// TIA Portal project "EbAndon v4_00_009" (V15) (continued)
DEVICE "ET 200SP station_27"  ET 200SP-Station
   slot 0: "Rack_0"  Rack  6ES5 710-8MAx1
   slot 0: "cv02et200sp"  IM 155-6 PN ST  6ES7 155-6AU01-0BN0  V4.1
   slot 1: "DQ 8x24VDC/0.5A ST_1"  DQ 8x24VDC/0.5A ST  6ES7 132-6BF01-0BA0  V0.0
      slot 1: "DQ 8x24VDC/0.5A ST_1"  DQ 8x24VDC/0.5A ST
   slot 2: "DQ 8x24VDC/0.5A ST_2"  DQ 8x24VDC/0.5A ST  6ES7 132-6BF01-0BA0  V0.0
      slot 1: "DQ 8x24VDC/0.5A ST_2"  DQ 8x24VDC/0.5A ST
   slot 3: "DQ 8x24VDC/0.5A ST_3"  DQ 8x24VDC/0.5A ST  6ES7 132-6BF01-0BA0  V0.0
      slot 1: "DQ 8x24VDC/0.5A ST_3"  DQ 8x24VDC/0.5A ST
   slot 4: "Server module_1"  Server module  6ES7 193-6PA00-0AA0  V1.1
      slot 1: "Server module_1"  Server module
   slot 127: "BA 2xRJ45"  BA 2xRJ45  6ES7 193-6AR00-0AA0  V0.0
      slot 1: "Port_1"  6ES7 193-6AR00-0AA0  V0.0
      slot 2: "Port_2"  6ES7 193-6AR00-0AA0  V0.0
DEVICE "ET 200SP station_28"  ET 200SP-Station
   slot 0: "Rack_0"  Rack  6ES5 710-8MAx1
   slot 0: "cv03et200sp"  IM 155-6 PN ST  6ES7 155-6AU01-0BN0  V4.1
   slot 1: "DQ 8x24VDC/0.5A ST_1"  DQ 8x24VDC/0.5A ST  6ES7 132-6BF01-0BA0  V0.0
      slot 1: "DQ 8x24VDC/0.5A ST_1"  DQ 8x24VDC/0.5A ST
   slot 2: "DQ 8x24VDC/0.5A ST_2"  DQ 8x24VDC/0.5A ST  6ES7 132-6BF01-0BA0  V0.0
      slot 1: "DQ 8x24VDC/0.5A ST_2"  DQ 8x24VDC/0.5A ST
   slot 3: "DQ 8x24VDC/0.5A ST_3"  DQ 8x24VDC/0.5A ST  6ES7 132-6BF01-0BA0  V0.0
      slot 1: "DQ 8x24VDC/0.5A ST_3"  DQ 8x24VDC/0.5A ST
   slot 4: "Server module_1"  Server module  6ES7 193-6PA00-0AA0  V1.1
      slot 1: "Server module_1"  Server module
   slot 127: "BA 2xRJ45"  BA 2xRJ45  6ES7 193-6AR00-0AA0  V0.0
      slot 1: "Port_1"  6ES7 193-6AR00-0AA0  V0.0
      slot 2: "Port_2"  6ES7 193-6AR00-0AA0  V0.0
DEVICE "ET 200SP station_29"  ET 200SP-Station
   slot 0: "Rack_0"  Rack  6ES5 710-8MAx1
   slot 0: "cv04et200sp"  IM 155-6 PN ST  6ES7 155-6AU01-0BN0  V4.1
   slot 1: "DQ 8x24VDC/0.5A ST_1"  DQ 8x24VDC/0.5A ST  6ES7 132-6BF01-0BA0  V0.0
      slot 1: "DQ 8x24VDC/0.5A ST_1"  DQ 8x24VDC/0.5A ST
   slot 2: "DQ 8x24VDC/0.5A ST_2"  DQ 8x24VDC/0.5A ST  6ES7 132-6BF01-0BA0  V0.0
      slot 1: "DQ 8x24VDC/0.5A ST_2"  DQ 8x24VDC/0.5A ST
   slot 3: "DQ 8x24VDC/0.5A ST_3"  DQ 8x24VDC/0.5A ST  6ES7 132-6BF01-0BA0  V0.0
      slot 1: "DQ 8x24VDC/0.5A ST_3"  DQ 8x24VDC/0.5A ST
   slot 4: "Server module_1"  Server module  6ES7 193-6PA00-0AA0  V1.1
      slot 1: "Server module_1"  Server module
   slot 127: "BA 2xRJ45"  BA 2xRJ45  6ES7 193-6AR00-0AA0  V0.0
      slot 1: "Port_1"  6ES7 193-6AR00-0AA0  V0.0
      slot 2: "Port_2"  6ES7 193-6AR00-0AA0  V0.0
DEVICE "ET 200SP station_30"  ET 200SP-Station
   slot 0: "Rack_0"  Rack  6ES5 710-8MAx1
   slot 0: "pc01et200sp"  IM 155-6 PN ST  6ES7 155-6AU01-0BN0  V4.1
   slot 1: "DQ 8x24VDC/0.5A ST_1"  DQ 8x24VDC/0.5A ST  6ES7 132-6BF01-0BA0  V0.0
      slot 1: "DQ 8x24VDC/0.5A ST_1"  DQ 8x24VDC/0.5A ST
   slot 2: "DQ 8x24VDC/0.5A ST_2"  DQ 8x24VDC/0.5A ST  6ES7 132-6BF01-0BA0  V0.0
      slot 1: "DQ 8x24VDC/0.5A ST_2"  DQ 8x24VDC/0.5A ST
   slot 3: "DQ 8x24VDC/0.5A ST_3"  DQ 8x24VDC/0.5A ST  6ES7 132-6BF01-0BA0  V0.0
      slot 1: "DQ 8x24VDC/0.5A ST_3"  DQ 8x24VDC/0.5A ST
   slot 4: "Server module_1"  Server module  6ES7 193-6PA00-0AA0  V1.1
      slot 1: "Server module_1"  Server module
   slot 127: "BA 2xRJ45"  BA 2xRJ45  6ES7 193-6AR00-0AA0  V0.0
      slot 1: "Port_1"  6ES7 193-6AR00-0AA0  V0.0
      slot 2: "Port_2"  6ES7 193-6AR00-0AA0  V0.0
DEVICE "ET 200SP station_31"  ET 200SP-Station
   slot 0: "Rack_0"  Rack  6ES5 710-8MAx1
   slot 0: "pc02et200sp"  IM 155-6 PN ST  6ES7 155-6AU01-0BN0  V4.1
   slot 1: "DQ 8x24VDC/0.5A ST_1"  DQ 8x24VDC/0.5A ST  6ES7 132-6BF01-0BA0  V0.0
      slot 1: "DQ 8x24VDC/0.5A ST_1"  DQ 8x24VDC/0.5A ST
   slot 2: "DQ 8x24VDC/0.5A ST_2"  DQ 8x24VDC/0.5A ST  6ES7 132-6BF01-0BA0  V0.0
      slot 1: "DQ 8x24VDC/0.5A ST_2"  DQ 8x24VDC/0.5A ST
   slot 3: "DQ 8x24VDC/0.5A ST_3"  DQ 8x24VDC/0.5A ST  6ES7 132-6BF01-0BA0  V0.0
      slot 1: "DQ 8x24VDC/0.5A ST_3"  DQ 8x24VDC/0.5A ST
   slot 4: "Server module_1"  Server module  6ES7 193-6PA00-0AA0  V1.1
      slot 1: "Server module_1"  Server module
   slot 127: "BA 2xRJ45"  BA 2xRJ45  6ES7 193-6AR00-0AA0  V0.0
      slot 1: "Port_1"  6ES7 193-6AR00-0AA0  V0.0
      slot 2: "Port_2"  6ES7 193-6AR00-0AA0  V0.0
*)

// ===== PLC "PLC_1"  CPU 1517F-3 PN/DP =====

VAR_GLOBAL   // PLC tag table "Default tag table"
   "System_Byte" AT %MB1 : Byte;
   "FirstScan" AT %M1.0 : Bool;
   "DiagStatUpdt" AT %M1.1 : Bool;
   "AlwaysTRUE" AT %M1.2 : Bool;
   "AlwaysFALSE" AT %M1.3 : Bool;
   "Clock_Byte" AT %MB0 : Byte;
   "Clock_10Hz" AT %M0.0 : Bool;
   "Clock_5Hz" AT %M0.1 : Bool;
   "Clock_2.5Hz" AT %M0.2 : Bool;
   "Clock_2Hz" AT %M0.3 : Bool;
   "Clock_1.25Hz" AT %M0.4 : Bool;
   "Clock_1Hz" AT %M0.5 : Bool;
   "Clock_0.625Hz" AT %M0.6 : Bool;
   "Clock_0.5Hz" AT %M0.7 : Bool;
   "Temp Reset" AT %M2.0 : Bool;
   "clearPartData" AT %M100.0 : Bool;
   "setDefaultPresets" AT %M100.1 : Bool;
   "hardInitReq" AT %M100.2 : Bool;
   "dbg" AT %M500.0 : Bool;
   "dbgSetDefTimes" AT %M5000.0 : Bool;
   "Copy PN Codes Into Recipes" AT %M10.0 : Bool;
   "Load Default Recipes Into Stations" AT %M10.1 : Bool;
   "Load Default Wip Data" AT %M10.2 : Bool;
   "dbg_station_index" AT %MW502 : Int;
END_VAR

VAR_GLOBAL CONSTANT   // PLC tag table "Default tag table"
   "ptsPerStn" : Int := 7;
   "slct_stn_btn_count" : Int := 11;
   "null_value" : Int := -1;
   "wip_pop_up_button_count" : Int := 6;   // number of wip select buttons on wip select pop up screen
END_VAR

VAR_GLOBAL   // PLC tag table "VOLVO 16 01"
   "VOLVO 16 01 IO" AT %QD1000 : DWord;
   "VOLVO 16 01 KP8 In" AT %ID0 : DWord;
   "VOLVO 16 01 KP8 Out" AT %QD0 : DWord;
END_VAR

VAR_GLOBAL   // PLC tag table "VOLVO 16 02"
   "VOLVO 16 02 IO" AT %QD1004 : DWord;
   "VOLVO 16 02 KP8 In" AT %ID4 : DWord;
   "VOLVO 16 02 KP8 Out" AT %QD4 : DWord;
END_VAR

VAR_GLOBAL   // PLC tag table "VOLVO 16 03"
   "VOLVO 16 03 IO" AT %QD1008 : DWord;
   "VOLVO 16 03 KP8 In" AT %ID8 : DWord;
   "VOLVO 16 03 KP8 Out" AT %QD8 : DWord;
END_VAR

VAR_GLOBAL   // PLC tag table "VOLVO 16 04"
   "VOLVO 16 04 IO" AT %QD1012 : DWord;
   "VOLVO 16 04 KP8 In" AT %ID12 : DWord;
   "VOLVO 16 04 KP8 Out" AT %QD12 : DWord;
END_VAR

VAR_GLOBAL   // PLC tag table "VOLVO 16 05"
   "VOLVO 16 05 IO" AT %QD1016 : DWord;
   "VOLVO 16 05 KP8 In" AT %ID16 : DWord;
   "VOLVO 16 05 KP8 Out" AT %QD16 : DWord;
END_VAR

VAR_GLOBAL   // PLC tag table "VOLVO 16 06"
   "VOLVO 16 06 IO" AT %QD1020 : DWord;
   "VOLVO 16 06 KP8 In" AT %ID20 : DWord;
   "VOLVO 16 06 KP8 Out" AT %QD20 : DWord;
END_VAR

VAR_GLOBAL   // PLC tag table "VOLVO 16 07"
   "VOLVO 16 07 IO" AT %QD1024 : DWord;
   "VOLVO 16 07 KP8 In" AT %ID24 : DWord;
   "VOLVO 16 07 KP8 Out" AT %QD24 : DWord;
END_VAR

VAR_GLOBAL   // PLC tag table "VOLVO 16 08"
   "VOLVO 16 08 IO" AT %QD1028 : DWord;
   "VOLVO 16 08 KP8 In" AT %ID28 : DWord;
   "VOLVO 16 08 KP8 Out" AT %QD28 : DWord;
END_VAR

VAR_GLOBAL   // PLC tag table "VOLVO 16 09"
   "VOLVO 16 09 IO" AT %QD1032 : DWord;
   "VOLVO 16 09 KP8 In" AT %ID32 : DWord;
   "VOLVO 16 09 KP8 Out" AT %QD32 : DWord;
END_VAR

VAR_GLOBAL   // PLC tag table "VOLVO 16 10"
   "VOLVO 16 10 IO" AT %QD1036 : DWord;
   "VOLVO 16 10 KP8 In" AT %ID36 : DWord;
   "VOLVO 16 10 KP8 Out" AT %QD36 : DWord;
END_VAR

VAR_GLOBAL   // PLC tag table "VOLVO 16 11"
   "VOLVO 16 11 IO" AT %QD1040 : DWord;
   "VOLVO 16 11 KP8 In" AT %ID40 : DWord;
   "VOLVO 16 11 KP8 Out" AT %QD40 : DWord;
END_VAR

VAR_GLOBAL   // PLC tag table "CHM 02"
   "CHM 02 KP8 In" AT %ID44 : DWord;
   "CHM 02 KP8 Out" AT %QD44 : DWord;
   "CHM 02 IO" AT %QD1044 : DWord;
END_VAR

VAR_GLOBAL   // PLC tag table "CHM 03"
   "CHM 03 IO" AT %QD1048 : DWord;
   "CHM 03 KP8 In" AT %ID48 : DWord;
   "CHM 03 KP8 Out" AT %QD48 : DWord;
END_VAR

VAR_GLOBAL   // PLC tag table "CHM 04"
   "CHM 04 IO" AT %QD1052 : DWord;
   "CHM 04 KP8 In" AT %ID52 : DWord;
   "CHM 04 KP8 Out" AT %QD52 : DWord;
END_VAR

VAR_GLOBAL   // PLC tag table "CHM 05"
   "CHM 05 IO" AT %QD1056 : DWord;
   "CHM 05 KP8 In" AT %ID56 : DWord;
   "CHM 05 KP8 Out" AT %QD56 : DWord;
END_VAR

VAR_GLOBAL   // PLC tag table "CDO 01"
   "CDO 01 IO" AT %QD1060 : DWord;
   "CDO 01 KP8 In" AT %ID60 : DWord;
   "CDO 01 KP8 Out" AT %QD60 : DWord;
END_VAR

VAR_GLOBAL   // PLC tag table "CDO 02"
   "CDO 02 IO" AT %QD1064 : DWord;
   "CDO 02 KP8 In" AT %ID64 : DWord;
   "CDO 02 KP8 Out" AT %QD64 : DWord;
END_VAR

VAR_GLOBAL   // PLC tag table "CDO 03"
   "CDO 03 IO" AT %QD1068 : DWord;
   "CDO 03 KP8 In" AT %ID68 : DWord;
   "CDO 03 KP8 Out" AT %QD68 : DWord;
END_VAR

VAR_GLOBAL   // PLC tag table "BFL 01"
   "BFL 01 IO" AT %QD1072 : DWord;
   "BFL 01 KP8 In" AT %ID72 : DWord;
   "BFL 01 KP8 Out" AT %QD72 : DWord;
   "Manual Operations Trigger" AT %M10.3 : Bool;
END_VAR

VAR_GLOBAL   // PLC tag table "BFL 02"
   "BFL 02 IO" AT %QD1076 : DWord;
   "BFL 02 KP8 In" AT %ID76 : DWord;
   "BFL 02 KP8 Out" AT %QD76 : DWord;
END_VAR

VAR_GLOBAL   // PLC tag table "BFL 03"
   "BFL 03 IO" AT %QD1080 : DWord;
   "BFL 03 KP8 In" AT %ID80 : DWord;
   "BFL 03 KP8 Out" AT %QD80 : DWord;
END_VAR

VAR_GLOBAL   // PLC tag table "LGS 01"
   "LGS 01 IO" AT %QD1084 : DWord;
   "LGS 01 KP8 In" AT %ID84 : DWord;
   "LGS 01 KP8 Out" AT %QD84 : DWord;
END_VAR

VAR_GLOBAL   // PLC tag table "LGS 02"
   "LGS 02 IO" AT %QD1088 : DWord;
   "LGS 02 KP8 In" AT %ID88 : DWord;
   "LGS 02 KP8 Out" AT %QD88 : DWord;
END_VAR

VAR_GLOBAL   // PLC tag table "CHM 01"
   "CHM 01 IO" AT %QD1092 : DWord;
   "CHM 01 KP8 In" AT %ID92 : DWord;
   "CHM 01 KP8 Out" AT %QD92 : DWord;
END_VAR

VAR_GLOBAL CONSTANT   // PLC tag table "Comm Diag"
   "pnioDeviceCount" : Int := 48;   // Upper limit of devices per HMI screen
   "USERDIAG_SLOTS_PER_SCREEN_UPPER_LIM" : Int := 31;   // Upper limit of slots per HMI screen
   "USERDIAG_SLOTS_PER_DEVICE_UPPER_LIM" : Int := 31;   // max number of modules per device
   "USERDIAG_DEVICES_PER_IO_SYSTEM_UPPER_LIM" : Int := 128;   // Upper limit of devices/slaves per IO-System/DP-Mastersystem
   "USERDIAG_SLOTS_PER_PLC_UPPER_LIM" : Int := 31;   // max number of local modules
   "USERDIAG_IO_SYSTEMS_UPPER_LIM" : Int := 1;   // Upper limit of IO-Systems/DP-Mastersystems
   "USERDIAG_IOSYSTEM_1" : Int := 1;   // Index for first IO-System/DP-Mastersystem
END_VAR

VAR_GLOBAL CONSTANT   // PLC tag table "Color Library"
   "BkBk" : USInt := 0;
   "BgWh" : USInt := 1;
   "FgWh" : USInt := 2;
   "FlWh" : USInt := 3;
   "BgGray" : USInt := 4;
   "FgGray" : USInt := 5;
   "FlGray" : USInt := 6;
   "BgLRd" : USInt := 7;
   "FgLRd" : USInt := 8;
   "FlLRd" : USInt := 9;
   "BgDRd" : USInt := 10;
   "FgDRd" : USInt := 11;
   "FlDrd" : USInt := 12;
   "BgLYe" : USInt := 13;
   "FgLYe" : USInt := 14;
   "FlLYe" : USInt := 15;
   "BgDYe" : USInt := 16;
   "FgDYe" : USInt := 17;
   "FlDYe" : USInt := 18;
   "BgLGr" : USInt := 19;
   "FgLGr" : USInt := 20;
   "FlLGr" : USInt := 21;
   "BgDGr" : USInt := 22;
   "FgDGr" : USInt := 23;
   "FlDGr" : USInt := 24;
   "BgLTe" : USInt := 25;
   "FgLTe" : USInt := 26;
   "FlLTe" : USInt := 27;
   "BgDTe" : USInt := 28;
   "FgDTe" : USInt := 29;
   "FlDTe" : USInt := 30;
   "BgLBl" : USInt := 31;
   "FgLBl" : USInt := 32;
   "FlLBl" : USInt := 33;
   "BgDBl" : USInt := 34;
   "FgDBl" : USInt := 35;
   "FlDBl" : USInt := 36;
   "BgLPu" : USInt := 37;
   "FgLPu" : USInt := 38;   // foreground light purple
   "FlLPu" : USInt := 39;
   "BgDPu" : USInt := 40;
   "FgDPu" : USInt := 41;
   "FlDPu" : USInt := 42;
   "disabled" : USInt := 254;
   "invisible" : USInt := 255;
   "LBlDRd" : USInt := 43;
   "DRdLBl" : USInt := 44;
   "LBlDRdFl" : USInt := 45;
   "DBlDRd" : USInt := 46;
   "DRdDBl" : USInt := 47;
   "DBlDRdFl" : USInt := 48;
END_VAR

VAR_GLOBAL CONSTANT   // PLC tag table "Station Meta Data"
   "btnCount" : Int := 7;   // one less than actual button count
   "stnCount" : Int := 38;   // one less than actual station count
   "defaultAlotted" : Real := 1800.0;
   "defaultCritical" : Real := 300.0;
   "wipCount" : Int := 49;   // one less than actual wip count
   "mStringLen" : Int := 40;
   "sStringLen" : Int := 20;
   "lStringLen" : Int := 100;
   "pnLibCount" : Int := 999;   // one less than actual pn capacity
   "kp8StnCount" : Int := 33;
   "hmi_station_count" : Int := 4;   // number of stations using basic panel instead of kp8 (-1 for array)
END_VAR

VAR_GLOBAL   // PLC tag table "Simulation"
   "simMode" AT %M100.3 : Bool;
END_VAR

VAR_GLOBAL CONSTANT   // PLC tag table "Simulation"
   "simKP8Count" : Int := 11;
END_VAR

VAR_GLOBAL CONSTANT   // PLC tag table "Station IDs"
   "VOLVO 16 01" : Int := 0;
   "VOLVO 16 02" : Int := 1;
   "VOLVO 16 03" : Int := 2;
   "VOLVO 16 04" : Int := 3;
   "VOLVO 16 05" : Int := 4;
   "VOLVO 16 06" : Int := 5;
   "VOLVO 16 07" : Int := 6;
   "VOLVO 16 08" : Int := 7;
   "VOLVO 16 09" : Int := 8;
   "VOLVO 16 10" : Int := 9;
   "VOLVO 16 11" : Int := 10;
   "CHM 01" : Int := 11;
   "CHM 02" : Int := 12;
   "CHM 03" : Int := 13;
   "CHM 04" : Int := 14;
   "CHM 05" : Int := 15;
   "CDO 01" : Int := 16;
   "CDO 02" : Int := 17;
   "CDO 03" : Int := 18;
   "BFL 01" : Int := 19;
   "BFL 02" : Int := 20;
   "BFL 03" : Int := 21;
   "LGS 01" : Int := 22;
   "LGS 02" : Int := 23;
   "LGS 03" : Int := 24;
   "CV 01" : Int := 25;
   "CV 02" : Int := 26;
   "CV 03" : Int := 27;
   "CV 04" : Int := 28;
   "PC 01" : Int := 29;
   "PC 02" : Int := 30;
END_VAR

VAR_GLOBAL CONSTANT   // PLC tag table "LED Sign"
   "ledRowCount" : Int := 11;
END_VAR

VAR_GLOBAL CONSTANT   // PLC tag table "HMI Part Request Screen"
   "partReqTblHMIRowCnt" : Int := 10;   // number of rows displayed on hmi
END_VAR

VAR_GLOBAL CONSTANT   // PLC tag table "HMI Settings Screen"
   "stngsScrnSlctdStns" : Int := 11;   // labels for settings screen
END_VAR

VAR_GLOBAL CONSTANT   // PLC tag table "Part Request Data Base"
   "partReqDataRowCount" : Int := 199;   // number of rows in part request table
END_VAR

VAR_GLOBAL CONSTANT   // PLC tag table "HMI Station"
   "wipSelScrnObjCnt" : Int := 29;   // number of buttons on menu select screen (short and long rows use different data, -1 for array)
   "partSelScrnObjCnt" : Int := 7;   // number of buttons on part select screen (-1 for array)
   "tmpltScrnObjCnt" : Int := 1;   // number of button on the template (-1 for array)
   "wip_select_button_count" : Int := 5;   // button count for wip selection screen on hmi stations, -1 for array
END_VAR

VAR_GLOBAL   // PLC tag table "LGS 03"
   "LGS 03 IO" AT %QD1096 : DWord;
   "LGS 03 KP8 In" AT %ID96 : DWord;
   "LGS 03 KP8 Out" AT %QD96 : DWord;
END_VAR

VAR_GLOBAL   // PLC tag table "CV 01"
   "CV 01 IO" AT %QD1100 : DWord;
   "CV 01 KP8 In" AT %ID100 : DWord;
   "CV 01 KP8 Out" AT %QD100 : DWord;
END_VAR

VAR_GLOBAL   // PLC tag table "CV 02"
   "CV 02 IO" AT %QD1104 : DWord;
   "CV 02 KP8 In" AT %ID104 : DWord;
   "CV 02 KP8 Out" AT %QD104 : DWord;
END_VAR

VAR_GLOBAL   // PLC tag table "CV 03"
   "CV 03 IO" AT %QD1108 : DWord;
   "CV 03 KP8 In" AT %ID108 : DWord;
   "CV 03 KP8 Out" AT %QD108 : DWord;
END_VAR

VAR_GLOBAL   // PLC tag table "CV 04"
   "CV 04 IO" AT %QD1112 : DWord;
   "CV 04 KP8 In" AT %ID112 : DWord;
   "CV 04 KP8 Out" AT %QD112 : DWord;
END_VAR

VAR_GLOBAL   // PLC tag table "PC 01"
   "PC 01 IO" AT %QD1116 : DWord;
   "PC 01 KP8 In" AT %ID116 : DWord;
   "PC 01 KP8 Out" AT %QD116 : DWord;
END_VAR

VAR_GLOBAL   // PLC tag table "PC 02"
   "PC 02 IO" AT %QD1120 : DWord;
   "PC 02 KP8 In" AT %ID120 : DWord;
   "PC 02 KP8 Out" AT %QD120 : DWord;
END_VAR

VAR_GLOBAL CONSTANT   // PLC tag table "States"
   "requested" : Int := 10;
   "ordered" : Int := 20;
   "requestedCrit" : Int := 11;
   "requestedExp" : Int := 12;
   "acknowledged" : Int := 30;
   "reset" : Int := 99;
   "idle" : Int := 01;
   "orderedCrit" : Int := 21;
   "acknowledgedCrit" : Int := 31;
   "orderedExp" : Int := 22;
   "acknowledgedExp" : Int := 32;
END_VAR

VAR_GLOBAL CONSTANT   // PLC tag table "Timers"
   "tCritical" : Real := 5.0;
   "tAllotted" : Real := 10.0;
END_VAR

TYPE "Station: All Stations"
   STRUCT
      stn : Array[0.."stnCount"] of "Station: Single Station";
   END_STRUCT;
END_TYPE

TYPE "Part Call Screen"
   STRUCT
      row : Array[0.."partReqTblHMIRowCnt"] of "Table Row";
   END_STRUCT;
END_TYPE

TYPE "Station: Wip: Wip Module"
   STRUCT
      ioData : "Station I/O Data";
      flags : "Station: Wip Flags";
      kp8Logical : "KP8 Driver: Feedback Data";
      orderState : Array[0.."btnCount"] of Int;
      pnCode : Array[0.."btnCount"] of DInt;
      timers : "Station: Timers";
      wip : "Station: Wip: Meta Data: Single";
   END_STRUCT;
END_TYPE

TYPE "Barcode Screen"
   STRUCT
      partNumber : WString[40];
      barcode : String;
      acknowledged : Bool;
      ordered : Bool;
   END_STRUCT;
END_TYPE

TYPE "Table Row"
   STRUCT
      address : DInt := -1;
      ordered : Bool;
      pbSelection : Struct
         actuate : Bool;
         animate : USInt;
      END_STRUCT;
      rtBackground : Struct
         animate : USInt;
      END_STRUCT;
      tfDropZone : Struct
         animate : USInt;
         value : WString[20];
      END_STRUCT;
      tfLine : Struct
         animate : USInt;
         value : WString[20];
      END_STRUCT;
      tfPartNumber : Struct
         animateDL : USInt;
         animateSL : USInt;
         value : WString[40];
      END_STRUCT;
      tfTime : Struct
         animate : USInt;
         value : WString[20];
      END_STRUCT;
   END_STRUCT;
END_TYPE

TYPE "Station: Order States"
   STRUCT
      btn : Array[0.."btnCount"] of Int;
   END_STRUCT;
END_TYPE

TYPE "Station: KP8 Config"
VERSION : 0.1
   STRUCT
      activate : Bool;
      colorOn1 : String[10];
      colorOn2 : String[10];
      colorOff : String[10];
      flash : Bool;
      group : Int;
      mode : Bool;
   END_STRUCT;
END_TYPE

TYPE "Station: PN Code"
   STRUCT
      btn : Array[0.."btnCount"] of DInt;
   END_STRUCT;
END_TYPE

TYPE "Part Request Data"
   STRUCT
      row : Array[0.."partReqDataRowCount"] of DInt;
   END_STRUCT;
END_TYPE

TYPE "Station: Single Station"
   STRUCT
      flags : "Station: Flags";
      id : "Station: Id";
      kp8Config : "KP8 Driver: Parameters: 8 Buttons";
      kp8Physical : "KP8 Driver: Feedback Data";
      wipData : "Station: Wip: Meta Data: All";
      wipCmpts : "Station: Wip: Wip Module";
   END_STRUCT;
END_TYPE

TYPE "Settings"
   STRUCT
      selectStation : "PB Data";
      selectWip : "PB Data";
      selectButton : "PB Data";
      line : "IO Field Data: Label with Data";
      dropzone : "IO Field Data: Label with Data";
      total : "IO Field Data: Label with Data";
      critical : "IO Field Data: Label with Data";
      partNumber : "IO Field Data: Label with Data";
      assign : "PB Data";
      stationRows : Array[0..2] of "Settings Station Row Data";
      stnTableNavBar : "Nav Bar Data: PLC";
   END_STRUCT;
   // selectStation.animate := 1;
END_TYPE

TYPE "PB Data"
   STRUCT
      actuate : Bool;
      animate : USInt;
      enable : Bool;
      label : WString[80];
      listSelect : UInt;
      visible : Bool;
   END_STRUCT;
END_TYPE

TYPE "LED Sign Data"
   STRUCT
      row : Array[0.."ledRowCount"] of "Table Row";
   END_STRUCT;
END_TYPE

TYPE "Nav Bar Data: HMI"
   STRUCT
      top_actuate : Bool;
      top_animate : USInt;
      top_enable : Bool;
      top_label : WString;
      top_list_select : UInt;
      top_visible : Bool;
      page_up_actuate : Bool;
      page_up_animate : USInt;
      page_up_enable : Bool;
      page_up_label : WString;
      page_up_list_select : UInt;
      page_up_visible : Bool;
      line_up_actuate : Bool;
      line_up_animate : USInt;
      line_up_enable : Bool;
      line_up_label : WString;
      line_up_list_select : UInt;
      line_up_visible : Bool;
      line_down_actuate : Bool;
      line_down_animate : USInt;
      line_down_enable : Bool;
      line_down_label : WString;
      line_down_list_select : UInt;
      line_down_visible : Bool;
      page_down_actuate : Bool;
      page_down_animate : USInt;
      page_down_enable : Bool;
      page_down_label : WString;
      page_down_list_select : UInt;
      page_down_visible : Bool;
      bottom_actuate : Bool;
      bottom_animate : USInt;
      bottom_enable : Bool;
      bottom_label : WString;
      bottom_list_select : UInt;
      bottom_visible : Bool;
   END_STRUCT;
END_TYPE

TYPE "Station: Animations"
   STRUCT
      btn : Array[0.."btnCount"] of UInt;
   END_STRUCT;
END_TYPE

TYPE "Pop Ups"
   STRUCT
      select_buttons : "Select Button";
      select_stations : "Select Station";
      select_WIPs : "Select WIP";
   END_STRUCT;
END_TYPE

TYPE "IO Field Data: Label with Data"
   STRUCT
      animate : USInt;
      enable : Bool;
      inputFinished : Bool;
      value : WString[40];
      visible : Bool;
   END_STRUCT;
END_TYPE

TYPE "Station Selection Change"
   STRUCT
      falling : Bool;
      rising : Bool;
      selection_change : Bool;
      station_index : Int := -1;
   END_STRUCT;
END_TYPE

TYPE "Selectable Station States"
   STRUCT
      all : Bool;
      non_hmi : Bool;
      hmi : Bool;
   END_STRUCT;
END_TYPE

TYPE "Selectable Stations"
   STRUCT
      stns : Array[0.."stnCount"] of Int;
   END_STRUCT;
END_TYPE

TYPE "Nav Bar Data: PLC"
   STRUCT
      top : "PB Data";
      pageUp : "PB Data";
      lineUp : "PB Data";
      lineDown : "PB Data";
      pageDown : "PB Data";
      bottom : "PB Data";
   END_STRUCT;
END_TYPE

TYPE "Station: Sim Data"
   STRUCT
      stn : Struct
         animate : USInt;
         label : WString[20];
      END_STRUCT;
      btn : Struct
         actuate : Byte;
         animate : Array[0..7] of USInt;
         labels : Array[0..7] of WString [4];
      END_STRUCT;
   END_STRUCT;
END_TYPE

TYPE "Simulated Stations"
   STRUCT
      down : "PB Data";
      firstStn : Int;
      me : Array[0.."simKP8Count"] of "Station: Sim Data";
      up : "PB Data";
   END_STRUCT;
END_TYPE

TYPE "Station: Wip Flags"
   STRUCT
      clearWipRequest : Bool;   // set: after wip has been deselected for deselect interval; consumed:
      inSettingsScreen : Bool;   // set: Flags: HMI Warehouse; consumed: Settings; reset: Flags: HMI Warehouse
      whHmiOrdered : Bool;   // set: Flags: HMI Warehouse, set by user input; consumed: Order State: Enter Ordered; reset: Order State: Enter Ordered
      newPN : Bool;   // set: Flags: New PN Code; reset:
      pnGood : Array[0.."btnCount"] of Bool;
      resetStation : Bool;
      resetTimer : Array[0.."btnCount"] of Bool;
   END_STRUCT;
END_TYPE

TYPE "HMI Station: Part Selection Screen"
   STRUCT
      animate : Array[0.."partSelScrnObjCnt"] of Int;
      pbs : DWord;
      txt : Array[0.."partSelScrnObjCnt"] of WString [40];
   END_STRUCT;
END_TYPE

TYPE "Runtime Data"
   STRUCT
      asReal : Real;
      elapsed : LReal;
      mem : LReal;
   END_STRUCT;
END_TYPE

TYPE "Recipe: Wip Text Library"
   STRUCT
      code : Array[0..99] of WString["sStringLen"];
      txt : Array[0..99] of WString["lStringLen"];
   END_STRUCT;
END_TYPE

TYPE "From Excel: Codes Single Wip"
VERSION : 0.1
   STRUCT
      pStn : Int := -1;
      pnCode : Array[0.."btnCount"] of DInt;
   END_STRUCT;
END_TYPE

TYPE "Recipe: HMI Stations Saved Wips"
   STRUCT
      stn : Array[0.."hmi_station_count"] of "WIP: Station";
   END_STRUCT;
END_TYPE

TYPE "Network Health Screen"
   STRUCT
      et200spPopUp : "Station: ET200SP Comm Debug Data";
      kp8PopUp : "Station: KP8 Comm Debug Data";
      pnioDevices : Array[1.."pnioDeviceCount"] of "PB Data";
      selectedDevice : Int;
   END_STRUCT;
END_TYPE

TYPE "HMI Stations"
   STRUCT
      stns : Array[0.."hmi_station_count"] of "HMI Station: Compressed";
   END_STRUCT;
END_TYPE

TYPE "Station: ET200SP Comm Debug Data"
   STRUCT
      dismissPB : Bool;
      IM : "ET200SP: IM Data";
      DQ01 : "ET200SP: DQ Data";
      DQ02 : "ET200SP: DQ Data";
      DQ03 : "ET200SP: DQ Data";
      profinetName : Struct
         animate : USInt;
         label : WString[20];
      END_STRUCT;
      serverModule : "ET200SP: Server Module Data";
   END_STRUCT;
END_TYPE

TYPE "ET200SP: IM Data"
   STRUCT
      bg : USInt;
      error : USInt;
      lnk01 : USInt;
      lnk02 : USInt;
      maint : USInt;
      pwr : USInt;
      run : USInt;
   END_STRUCT;
END_TYPE

TYPE "ET200SP: DQ Data"
   STRUCT
      bg : USInt;
      bgTem : USInt;
      diag : USInt;
      pwr : USInt;
      x0 : USInt;
      x1 : USInt;
      x2 : USInt;
      x3 : USInt;
      x4 : USInt;
      x5 : USInt;
      x6 : USInt;
      x7 : USInt;
   END_STRUCT;
END_TYPE

TYPE "ET200SP: Server Module Data"
   STRUCT
      bg : USInt;
   END_STRUCT;
END_TYPE

TYPE "Station: KP8 Comm Debug Data"
   STRUCT
      dismissPB : Bool;
      profinetName : Struct
         animate : USInt;
         label : WString[20];
      END_STRUCT;
      stencilBackground : USInt;
      X1P1 : Struct
         transmit : USInt;
         receive : USInt;
      END_STRUCT;
      X1P2 : Struct
         transmit : USInt;
         receive : USInt;
      END_STRUCT;
   END_STRUCT;
END_TYPE

TYPE "From Excel: Codes Multiple Wips"
VERSION : 0.1
   STRUCT
      pStn : Int := -1;
      wip : Array[0.."wipCount"] of Struct
         wipCode : DInt;
         pnCode : Array[0.."btnCount"] of DInt;
      END_STRUCT;
   END_STRUCT;
END_TYPE

TYPE "Station: Timers"
   STRUCT
      elapsed : Array[0.."btnCount"] of Real;   // time (s) that a part number has been requested
      ptAllotted : Array[0.."btnCount"] of Real;   // time (s) before a part request is considered over-due
      ptCritical : Array[0.."btnCount"] of Real;   // time (s) before a part request is considered critical
      remaining : Array[0.."btnCount"] of Real;   // request allotted - elapsed
      wsAllotted : Real := 10.0;   // time (s) before a selected wip is counted as being selected
      wsElapsed : Real;   // time (s) a wip has been selected
      wsRemaining : Real;   // wip select allotted - selected
      wdsAllotted : Real := 10.0;   // time (s) before a deselected wip's requests are cleared from the part request table
      wdsElapsed : Real;   // time (s) a wip has been deselected
      wdsRemaining : Real;   // wip deselect allotted - selected
   END_STRUCT;
END_TYPE

TYPE "Station: Wip: Meta Data: Single"
   STRUCT
      code : DInt := -1;   // builds station name from libraries
      useCount : DInt;   // number of times station selected for longer than lower dwell limit
   END_STRUCT;
END_TYPE

TYPE "HMI Station: Wip Select: PLC Interface"
   STRUCT
      raw : Array[0..31] of Bool;
      wsRising : Array[0..5] of Bool;
      wsFalling : Array[0..5] of Bool;
   END_STRUCT;
END_TYPE

TYPE "Settings Station Row Data"
   STRUCT
      line : "Cell Data";
      dropzone : "Cell Data";
      wip : "Cell Data";
      btnRows : Array[0..7] of "Settings Station Row Button Row Data";
   END_STRUCT;
END_TYPE

TYPE "Station: Flags"
   STRUCT
      stateTransition : Array[0.."btnCount"] of Bool;
      wipSwapped : Bool;
   END_STRUCT;
END_TYPE

TYPE "HMI Station: Compressed"
   STRUCT
      partSelect : "HMI Station: Part Selection Screen";
      template : "HMI Station: Template Screen";
      wipSelect : "HMI Station: Wip Select: Screen";
   END_STRUCT;
END_TYPE

TYPE "HMI Station: Wip Select: Screen"
   STRUCT
      animate : Array[0.."wipSelScrnObjCnt"] of Int;
      pbs : DWord;
      txt : Array[0.."wipSelScrnObjCnt"] of WString ["lStringLen"];
   END_STRUCT;
   // // txt[6] : wip select 00 label
   // // txt[7] : wip select 00 text
   // // txt[8] : wip select 01 label
   // // txt[9] : wip select 01 text
   // // txt[10] : wip select 02 label
   // // txt[11] : wip select 02 text
   // // txt[12] : wip select 03 label
   // // txt[13] : wip select 03 text
   // // txt[14] : wip select 04 label
   // // txt[15] : wip select 04 text
   // // txt[16] : wip select 05 label
   // // txt[17] : wip select 05 text
END_TYPE

TYPE "HMI Station: Template Screen"
   STRUCT
      animate : Array[0.."tmpltScrnObjCnt"] of Int;
      pb : DWord;
      text : Array[0.."tmpltScrnObjCnt"] of WString ["lStringLen"];
   END_STRUCT;
END_TYPE

TYPE "Selected Stations"
   STRUCT
      stns : Array[0.."stnCount"] of Bool;
   END_STRUCT;
END_TYPE

TYPE "Station: Id"
   STRUCT
      dropZone : USInt;
      lineName : WString["sStringLen"];
   END_STRUCT;
END_TYPE

TYPE "KP8 I/O Data"
   STRUCT
      input : Word;
      tempOut : DWord;
      finalOut : DWord;
   END_STRUCT;
END_TYPE

TYPE "Station I/O Data"
   STRUCT
      kp8 : "KP8 I/O Data";
      stkLight : DWord;
   END_STRUCT;
END_TYPE

